// Mitsubishi GX Works2 project: ZhaoQing_OCV__Debug   PLC: Q10UDEH (continued)
     
     (*空框换内衬线体*)
    SwitchIO12203.xEntryEnable:=  ConveyorIO12125.xNextRun;
    ConveyorIO12142.iProductCategoryIn:=ConveyorIO12125.iProductCategoryOut;
    IF ConveyorIO12142.iProductCategory=4 THEN
    	SwitchIO12203.xSwithEnable:=1;
    ELSE
    	SwitchIO12203.xSwithEnable:=0;
    END_IF;
    SwitchIO12203.xExitEnable:=ConveyorIO12143.xEmpty;
    ConveyorIO12143.xLoad:=ConveyorIO12142.xNextRun;
    ConveyorIO12143.iProductCategoryIn:=ConveyorIO12142.iProductCategoryOut;
    ConveyorIO12143.xUnload:=ConveyorIO12144.xEmpty;
    (*OCV1线体*) 
  (*  ConveyorIO12144.xLoad:=ConveyorIO12143.xNextRun;*)
    SwitchIO12330.xEntryEnable:=ConveyorIO12143.xNextRun;
    ConveyorIO12144.iProductCategoryIn:=ConveyorIO12143.iProductCategoryOut;
    IF ConveyorIO12144.iProductCategory =2 THEN  (*临时程序  手动调试完毕后改为2*)
   	 SwitchIO12330.xSwithEnable:=1;
    ELSE
    SwitchIO12330.xSwithEnable:=0;	
    END_IF;   
    ConveyorIO12144.xUnload:=ConveyorIO12333.xEmpty AND SwitchIO12330.xSwithEnable=0;
     SwitchIO12330.xExitEnable:=ConveyorIO12160.xEmpty AND SwitchIO12330.xSwithEnable=1;
     ConveyorIO12160.xLoad:=Switch12330ConveyorOut.xNextRun;
     IF XA5 THEN(*人工按钮*)
     	IF ConveyorIO12146.xEmpty THEN
     		m_xOCV1Done:=1;
     	END_IF;
     	m_xPickOutDone :=1;
     END_IF;
     IF ConveyorIO12160.xEmpty THEN
     	m_xOCV1Done:=0;
     END_IF ;
     IF ConveyorIO12146.xEmpty THEN
     	m_xPickOutDone :=0;
     END_IF;
     ConveyorIO12160.tLoadDelay:=T#2s;
     ConveyorIO12160.xUnload:=ConveyorIO12146.xEmpty AND m_xOCV1Done;
     Y27F:=ConveyorIO12146.xEmpty AND m_xOCV1Done;(*阻挡气缸*)
     ConveyorIO12146.xLoad:= ConveyorIO12160.xNextRun;
     (*OCV2线体*)    
    SwitchIO12333.xEntryEnable:=ConveyorIO12144.xNextRun;
	SwitchIO12333.xSwithEnable:=1;
	SwitchIO12333.xExitEnable:=NOT XAE;
     (*空框换内衬线体*)    	
     SwitchIO12204.xEntryEnable:=1;
      SwitchIO12204.xSwithEnable:=1;
      SwitchIO12204.xExitEnable:=ConveyorIO12151.xEmpty;
      ConveyorIO12151.xLoad:=ConveyorIO12204.xNextRun;
      ConveyorIO12151.xUnload:=ConveyorIO12150.xEmpty;
      ConveyorIO12150.xLoad:=ConveyorIO12151.xNextRun;
      ConveyorIO12150.xUnload:=ConveyorIO12149.xEmpty;
      SwitchIO12328.xEntryEnable:=ConveyorIO12150.xNextRun;
       SwitchIO12328.xSwithEnable:=1;
	(****************提升机8******************)
	Lifter8Priority(xCondition1:= NOT ConveyorIO12148.xEmpty,
	                          xCondition2:= NOT ConveyorIO12146.xEmpty AND m_xPickOutDone  ,
	                          xCondition3:= FALSE,(*成品库车间空框回流线体不为空的条件*)
	                          xCondition4:= FALSE ,
	                          xCondition5:= FALSE ,
	                          xTaskComplete:= LDF(TRUE,Conveyor8IO.xEmpty=0) ,
	                          xReset:=g_xResetSingle AND g_iDeviceIDSelect=8,
	                          iPriority:= m_iLifter8Task);
	     D16:=m_iLifter8Task;(*触摸屏显示当前任务*)
		CASE m_iLifter8Task OF
			1:(*空框回流线体*)
				Lifter8IO.iDestinationPos:=2;
				SwitchIO12328.xExitEnable:=Lifter8IO.iCurrentPos=2 AND XC2 AND Conveyor8IO.xEmpty AND NOT XC1;
			   Conveyor8IO.xLoad:=ConveyorIO12148.xNextRun;
               Conveyor8IO.xloadCCW:=1;
			2:(*OCV1*)
				Lifter8IO.iDestinationPos:=1;
			   Conveyor8IO.xLoad:=ConveyorIO12146.xNextRun;
			   ConveyorIO12146.xUnload:=Conveyor8Io.xEmpty AND Lifter8IO.iCurrentPos=1 AND XC1 AND XC2;
			   Y27E:=Conveyor8Io.xEmpty AND Lifter8IO.iCurrentPos=1 AND XC1 AND XC2;(*分拣位置阻挡气缸*)
               Conveyor8IO.xloadCCW:=0;			
			3:(*成品库对接*)
				Lifter8IO.iDestinationPos:=4;
			(*	Conveyor8IO.xLoad:=ConveyorIO12147.xNextRun;*)
				Conveyor8IO.xloadCCW:=0;
				ELSE
				Conveyor8IO.xLoad:=0;
				SwitchIO12328.xExitEnable:=0;
				ConveyorIO12146.xUnload:=0;
				Y27E:=0;(*分拣位置阻挡气缸*)
		END_CASE;		
	IF Conveyor8IO.xEmpty=0 THEN
		Lifter8IO.xMDIExe:=1;
		Lifter8IO.iDestinationPos:=3;
	END_IF;	
	IF Lifter8IO.iCurrentPos=3 AND XC3 THEN
		Conveyor8Io.xUnload:=ConveyorIO12159.xEmpty;
		Conveyor8IO.xUnloadCCW:=1;
	ELSE
		Conveyor8Io.xUnload:=0;
	END_IF;	
	ConveyorIO12159.xLoad:=Conveyor8IO.xNextRun;
   ConveyorIO12159.xUnload:=ConveyorIO12158.xEmpty;
   SwitchIO12337.xEntryEnable:=ConveyorIO12159.xNextRun;
   SwitchIO12337.xSwithEnable:=1;
   SwitchIO12337.xLiftCylinderExtendInit:=1;
   SwitchIO12337.xExitEnable:=ConveyorIO12156.xEmpty;
   ConveyorIO12156.xLoad:=ConveyorIO12157.xNextRun;
	(**********常温库入库分流*******************)	
	ConveyorIO12156.xUnload:=ConveyorIO12155.xEmpty;
	ConveyorIO12155.xLoad:=ConveyorIO12156.xNextRun;
	     (*触摸屏上计数与清零程序*)
     IF LDF(TRUE,ConveyorIO12155.xEmpty) THEN
     	D14:=D14+1;
     END_IF;
     IF M169 THEN
     	D14:=0;
     END_IF;
	
	(**********常温库1巷道入库*******************) 
         	ConveyorIO12155.xUnload:=ConveyorIO12141.xEmpty AND ConveyorIO12155.iProductCategory>1 ;
         	ConveyorIO12141.xLoad:=ConveyorIO12155.xNextRun;
         	ConveyorIO12141.xUnload:=ConveyorIO12321.xEmpty;
            (*分流信息传递到巷道1的顶升移载处*)        	
  			ConveyorIO12141.iProductCategoryIn:= ConveyorIO12155.iProductCategoryOut;    
  			    
            SwitchIO12321.xEntryEnable:=ConveyorIO12141.xNextRun;
			ConveyorIO12321.iProductCategoryIn:=ConveyorIO12141.iProductCategoryOut;
           (*分流信息显示为本巷道，启动顶升移载*)
           IF ConveyorIO12321.iProductCategory=2 THEN
          	 SwitchIO12321.xSwithEnable:=1;
           ELSE
      	     	SwitchIO12321.xSwithEnable:=0;
           END_IF;
           (*双料入库，优先选择1 ，当1结束后恢复到0，2秒 ，然后再跳到2,0状态用来复位移载的出料*) 
          m_tonSwitch1NOSeleteDelay(IN:= m_iSwitch12321Select=0 ,PT:= t#2S ,Q:=m_xSwitch12321NoSeleteDelay,ET:= m_tSwitch12321NOSeleteCurrent);
         IF   m_xSwitch12321NoSeleteDelay THEN
         	m_xSwitch12321Select:=1;
         END_IF;
         IF ldf(TRUE,ConveyorIO12138.xEmpty)  OR ldf(TRUE,ConveyorIO12139.xEmpty) THEN
         	m_xSwitch12321Select:=0;
         END_IF;
           IF ConveyorIO12139.xEmpty AND  m_xSwitch12321Select  THEN
           		m_iSwitch12321Select:=1;
	           	ELSIF NOT ConveyorIO12139.xEmpty  AND ConveyorIO12138.xEmpty AND m_xSwitch12321Select THEN
           	  	m_iSwitch12321Select:=2;
          	 ELSE
           		m_iSwitch12321Select:=0;
           END_IF;
           IF SwitchIO12321.xSwithEnable THEN
         	  SwitchIO12321.xExitEnable:=((ConveyorIO12139.xEmpty AND m_iSwitch12321Select=1) 
                                                          OR   (ConveyorIO12138.xEmpty AND m_iSwitch12321Select=2)) AND CylinderIO12320.iCurrentPos=1;
           ELSE(*分流到下一巷道*)
   	        	 SwitchIO12321.xExitEnable:= ConveyorIO12137.xEmpty;
    	        ConveyorIO12137.xLoad:= ConveyorIO12321.xNextRun ;
    	         ConveyorIO12137.iProductCategoryIn:=   ConveyorIO12321.iProductCategoryOut;     
            END_IF;
 
           ConveyorIO12139.xLoad:=ConveyorIO12140.xNextRun AND m_iSwitch12321Select=1 ;
   	       ConveyorIO12138.xLoad:=ConveyorIO12140.xNextRun AND m_iSwitch12321Select=2 ;
   	       IF  ConveyorIO12138.xEmpty =0 AND ConveyorIO12139.xEmpty =0 AND X72 AND X74 THEN
   	       	CylinderIO12320.xMDIExe:=1;
   	       	CylinderIO12320.iDestinationPos:=2;
   	       	ConveyorIO12138.xPutInto:=0;
   	       	ConveyorIO12139.xPutInto:=0;
   	       END_IF;
   	       IF g_xImport1Force THEN (* 1巷道单框强制入库*)
   	       	CylinderIO12320.xMDIExe:=1;
   	       	CylinderIO12320.iDestinationPos:=2;
   	       	ConveyorIO12138.xPutInto:=0;
   	       	ConveyorIO12139.xPutInto:=0;   
   	       	END_IF;	       
   	       IF NOT X72 AND NOT X74 THEN
   	       		CylinderIO12320.xMDIExe:=1;
   	       		CylinderIO12320.iDestinationPos:=1;
   	       END_IF;
   	       IF LDP(TRUE,CylinderIO12320.iCurrentPos=1 AND NOT ConveyorIO12138.xCWPresent AND NOT ConveyorIO12139.xCWPresent) THEN   	       	
   	       		ConveyorIO12138.xPutInto:=1;
   	       		ConveyorIO12139.xPutInto:=1;
   	       END_IF;        
	(**********常温库2巷道入库*******************)
	       ConveyorIO12137.xUnload:=ConveyorIO12136.xEmpty;
	       ConveyorIO12136.xLoad:=ConveyorIO12137.xNextRun;	       
  		   ConveyorIO12136.iProductCategoryIn:= ConveyorIO12137.iProductCategoryOut;  
         	ConveyorIO12136.xUnload:=ConveyorIO12135.xEmpty AND ConveyorIO12136.iProductCategory>2 ;
            (*分流信息传递到巷道1的顶升移载处*)        	
  			ConveyorIO12135.iProductCategoryIn:= ConveyorIO12136.iProductCategoryOut;       			    
            SwitchIO12317.xEntryEnable:=ConveyorIO12136.xNextRun;
           (*分流信息显示为本巷道，启动顶升移载*)
           IF ConveyorIO12135.iProductCategory=3 THEN
          	 SwitchIO12317.xSwithEnable:=1;
           ELSE
      	     	SwitchIO12317.xSwithEnable:=0;
           END_IF;
           (*双料入库，优先选择1 ，当1结束后恢复到0，2秒 ，然后再跳到2,0状态用来复位移载的出料*) 
          m_tonSwitch2NOSeleteDelay(IN:= m_iSwitch12317Select=0 ,PT:= t#2S ,Q:=m_xSwitch12317NoSeleteDelay,ET:= m_tSwitch12317NOSeleteCurrent);
         IF   m_xSwitch12317NoSeleteDelay THEN
         	m_xSwitch12317Select:=1;
         END_IF;
         IF ldf(TRUE,ConveyorIO12132.xEmpty)  OR ldf(TRUE,ConveyorIO12133.xEmpty) THEN
         	m_xSwitch12317Select:=0;
         END_IF;
           IF ConveyorIO12133.xEmpty AND  m_xSwitch12317Select   THEN
           		m_iSwitch12317Select:=1;
	           	ELSIF NOT ConveyorIO12133.xEmpty  AND ConveyorIO12132.xEmpty AND m_xSwitch12317Select THEN
           	  	m_iSwitch12317Select:=2;
          	 ELSE
           		m_iSwitch12317Select:=0;
           END_IF;
           IF SwitchIO12317.xSwithEnable THEN
         	  SwitchIO12317.xExitEnable:=((ConveyorIO12133.xEmpty AND m_iSwitch12317Select=1) 
                                                          OR   (ConveyorIO12132.xEmpty AND m_iSwitch12317Select=2)) AND CylinderIO12316.iCurrentPos=1;
           ELSE(*分流到下一巷道*)
   	        	 SwitchIO12317.xExitEnable:= ConveyorIO12131.xEmpty;
    	        ConveyorIO12131.xLoad:= ConveyorIO12135.xNextRun ;
    	        ConveyorIO12131.iProductCategoryIn:=ConveyorIO12135.iProductCategoryOut;
            END_IF;
           	                                          
           ConveyorIO12133.xLoad:=ConveyorIO12134.xNextRun AND m_iSwitch12317Select=1 ;
   	       ConveyorIO12132.xLoad:=ConveyorIO12134.xNextRun AND m_iSwitch12317Select=2 ;
   	       IF  ConveyorIO12133.xEmpty =0 AND ConveyorIO12132.xEmpty =0 AND CylinderIO12316.xPresentDetect1 AND CylinderIO12316.xPresentDetect2 THEN
   	       	CylinderIO12316.xMDIExe:=1;
   	       	CylinderIO12316.iDestinationPos:=2;
   	       	ConveyorIO12133.xPutInto:=0;
   	       	ConveyorIO12132.xPutInto:=0;
   	       END_IF;
   	       IF g_xImport2Force THEN (* 1巷道单框强制入库*)
   	       	CylinderIO12316.xMDIExe:=1;
   	       	CylinderIO12316.iDestinationPos:=2;
   	       	ConveyorIO12133.xPutInto:=0;
   	       	ConveyorIO12132.xPutInto:=0;   
   	       	END_IF;	       
   	       IF NOT CylinderIO12316.xPresentDetect1 AND NOT CylinderIO12316.xPresentDetect2 THEN
   	       		CylinderIO12316.xMDIExe:=1;
   	       		CylinderIO12316.iDestinationPos:=1;
   	       END_IF;
   	       IF LDP(TRUE,CylinderIO12316.iCurrentPos=1 AND NOT ConveyorIO12132.xCWPresent AND NOT ConveyorIO12133.xCWPresent) THEN   	       	
   	       		ConveyorIO12133.xPutInto:=1;
   	       		ConveyorIO12132.xPutInto:=1;
   	       END_IF;  
	(**********常温库3巷道入库*******************)
	       ConveyorIO12131.xUnload:=ConveyorIO12130.xEmpty AND ConveyorIO12131.iProductCategory>3 ;
	       ConveyorIO12130.xLoad:=ConveyorIO12131.xNextRun;	       
  		   ConveyorIO12130.iProductCategoryIn:= ConveyorIO12131.iProductCategoryOut;  
            (*分流信息传递到巷道1的顶升移载处*)   
             ConveyorIO12130.xUnload:=ConveyorIO12129.xEmpty;
             SwitchIO12314.xEntryEnable:=ConveyorIO12130.xNextRun;   	
  			ConveyorIO12129.iProductCategoryIn:= ConveyorIO12130.iProductCategoryOut;       			               
           (*分流信息显示为本巷道，启动顶升移载*)
           IF ConveyorIO12129.iProductCategory=4THEN
          	 SwitchIO12314.xSwithEnable:=1;
           ELSE
      	     	SwitchIO12314.xSwithEnable:=0;
           END_IF;
           (*双料入库，优先选择1 ，当1结束后恢复到0，2秒 ，然后再跳到2,0状态用来复位移载的出料*) 
          m_tonSwitch3NOSeleteDelay(IN:= m_iSwitch12314Select=0 ,PT:= t#2S ,Q:=m_xSwitch12314NoSeleteDelay,ET:= m_tSwitch12314NOSeleteCurrent);
         IF   m_xSwitch12314NoSeleteDelay THEN
         	m_xSwitch12314Select:=1;
         END_IF;
         IF ldf(TRUE,ConveyorIO12126.xEmpty)  OR ldf(TRUE,ConveyorIO12127.xEmpty) THEN
         	m_xSwitch12314Select:=0;
         END_IF;
           IF ConveyorIO12127.xEmpty AND  m_xSwitch12314Select   THEN
           		m_iSwitch12314Select:=1;
	           	ELSIF NOT ConveyorIO12127.xEmpty  AND ConveyorIO12126.xEmpty AND m_xSwitch12314Select THEN
           	  	m_iSwitch12314Select:=2;
          	 ELSE
           		m_iSwitch12314Select:=0;
           END_IF;
           IF SwitchIO12314.xSwithEnable THEN
         	  SwitchIO12314.xExitEnable:=((ConveyorIO12127.xEmpty AND m_iSwitch12314Select=1) 
                                                          OR   (ConveyorIO12126.xEmpty AND m_iSwitch12314Select=2)) AND CylinderIO12313.iCurrentPos=1;
           ELSE(*分流到下一巷道*)
				;(*报警*)
            END_IF;
           	                                          
           ConveyorIO12127.xLoad:=ConveyorIO12128.xNextRun AND m_iSwitch12314Select=1 ;
   	       ConveyorIO12126.xLoad:=ConveyorIO12128.xNextRun AND m_iSwitch12314Select=2 ;
   	       IF  ConveyorIO12126.xEmpty =0 AND ConveyorIO12127.xEmpty =0 AND CylinderIO12313.xPresentDetect1 AND CylinderIO12313.xPresentDetect2 THEN
   	       	CylinderIO12313.xMDIExe:=1;
   	       	CylinderIO12313.iDestinationPos:=2;
   	       	ConveyorIO12126.xPutInto:=0;
   	       	ConveyorIO12127.xPutInto:=0;
   	       END_IF;
   	       IF g_xImport3Force THEN (* 1巷道单框强制入库*)
   	       	CylinderIO12313.xMDIExe:=1;
   	       	CylinderIO12313.iDestinationPos:=2;
   	       	ConveyorIO12126.xPutInto:=0;
   	       	ConveyorIO12127.xPutInto:=0;   
   	       	END_IF;	       
   	       IF NOT CylinderIO12313.xPresentDetect1 AND NOT CylinderIO12313.xPresentDetect2 THEN
   	       		CylinderIO12313.xMDIExe:=1;
   	       		CylinderIO12313.iDestinationPos:=1;
   	       END_IF;
   	       IF LDP(TRUE,CylinderIO12313.iCurrentPos=1 AND NOT ConveyorIO12127.xCWPresent AND NOT ConveyorIO12126.xCWPresent) THEN   	       	
   	       		ConveyorIO12126.xPutInto:=1;
   	       		ConveyorIO12127.xPutInto:=1;
   	       END_IF;  
END_IF;
(*人工操作按钮*)
IF LDP(TRUE,X0FF)  AND NOT  Y290 THEN
	 m_xMotorFlag:=1;
ELSE
	m_xMotorFlag:=0;
END_IF;

IF m_xMotorFlag THEN
	Y290:=1;
	Y27A:=1;
	Y27B:=1;
END_IF;

IF LDP(TRUE,X0FF) AND NOT m_xMotorFlag THEN
	Y290:=0;
	Y27A:=0;
	Y27B:=0;
END_IF;
(*报警*)
M500:=D2330=1;(*常温库出库分流读码失败*)
M501:=D2325=1;(*常温库入库分流读码失败*)
g_xAlarm:=M500 
                     OR M501;
END_PROGRAM

FUNCTION_BLOCK PriorityFB
VAR_INPUT
  xCondition1 : BOOL;  (* 条件1 *)
  xCondition2 : BOOL;  (* 条件2 *)
  xCondition3 : BOOL;  (* 条件3 *)
  xCondition4 : BOOL;  (* 条件4 *)
  xCondition5 : BOOL;  (* 条件5 *)
  xTaskComplete : BOOL;  (* 任务完成 *)
  xReset : BOOL;  (* 复位 *)
END_VAR
VAR
  xOccupy : BOOL;  (* 占用 *)
END_VAR
VAR_OUTPUT
  iPriority : INT;  (* 输出任务号 *)
END_VAR
VAR
  m_tonCondition1Delay : TON;
  m_xCondition1Delay : BOOL;
  m_tCondition1CurrentTime : TIME;
  arriTaskStack : ARRAY [0..5] OF INT;
  m_tonCondition2Delay : TON;
  m_xCondition2Delay : BOOL;
  m_tCondition2CurrentTime : TIME;
  m_tonCondition3Delay : TON;
  m_xCondition3Delay : BOOL;
  m_tCondition3CurrentTime : TIME;
  m_tonCondition4Delay : TON;
  m_xCondition4Delay : BOOL;
  m_tCondition4CurrentTime : TIME;
  m_tonCondition5Delay : TON;
  m_xCondition5Delay : BOOL;
  m_tCondition5CurrentTime : TIME;
  jj : INT;
END_VAR
(****************************************************************************)
(*
优先级功能块，存储5个条件的优先级，实现栈功能先入先出，
复位功能还有问题，
*)
(***************************************************************************)
m_tonCondition1Delay(IN:= xCondition1 AND NOT xReset ,PT:= T#1s,Q:= m_xCondition1Delay , ET:= m_tCondition1CurrentTime );
m_tonCondition2Delay(IN:= xCondition2 AND NOT xReset ,PT:= T#1s,Q:= m_xCondition2Delay , ET:= m_tCondition2CurrentTime );
m_tonCondition3Delay(IN:= xCondition3 AND NOT xReset ,PT:= T#1s,Q:= m_xCondition3Delay , ET:= m_tCondition3CurrentTime );
m_tonCondition4Delay(IN:= xCondition4 AND NOT xReset ,PT:= T#1s,Q:= m_xCondition4Delay , ET:= m_tCondition4CurrentTime );
m_tonCondition5Delay(IN:= xCondition5 AND NOT xReset ,PT:= T#1s,Q:= m_xCondition5Delay , ET:= m_tCondition5CurrentTime );

IF ldp(TRUE,m_xCondition1Delay) THEN
	FOR jj:=0 TO 5 BY 1 DO
		IF arriTaskStack[jj]=0 THEN
			arriTaskStack[jj]:=1;
			EXIT;
		END_IF;		
	END_FOR;
END_IF;

IF ldp(TRUE,m_xCondition2Delay) THEN
	FOR jj:=0 TO 5 BY 1 DO
		IF arriTaskStack[jj]=0 THEN
			arriTaskStack[jj]:=2;
			EXIT;
		END_IF;		
	END_FOR;
END_IF;

IF ldp(TRUE,m_xCondition3Delay) THEN
	FOR jj:=0 TO 5 BY 1 DO
		IF arriTaskStack[jj]=0 THEN
			arriTaskStack[jj]:=3;
			EXIT;
		END_IF;		
	END_FOR;
END_IF;

IF ldp(TRUE,m_xCondition4Delay) THEN
	FOR jj:=0 TO 5 BY 1 DO
		IF arriTaskStack[jj]=0 THEN
			arriTaskStack[jj]:=4;
			EXIT;
		END_IF;		
	END_FOR;
END_IF;

IF ldp(TRUE,m_xCondition5Delay) THEN
	FOR jj:=0 TO 5 BY 1 DO
		IF arriTaskStack[jj]=0 THEN
			arriTaskStack[jj]:=5;
			EXIT;
		END_IF;		
	END_FOR;
END_IF;

iPriority:=arriTaskStack[0];

IF 	LDP(TRUE, xTaskComplete) THEN
	FOR jj:=0 TO 4 BY 1 DO
		arriTaskStack[jj]:=arriTaskStack[jj+1];
	END_FOR;
		arriTaskStack[5]:=0;
END_IF;

IF LDP(TRUE,xReset) THEN
		FOR jj:=0 TO 5 BY 1 DO
		arriTaskStack[jj]:=0;
	END_FOR;
END_IF;
END_FUNCTION_BLOCK

FUNCTION ShuttleCarCurrentPosition
VAR_INPUT
  xPosition1 : BOOL;
  xPosition2 : BOOL;
  xPosition3 : BOOL;
END_VAR
(************************************
计算输送车当前位置的函数
**************************************)
IF xPosition1 THEN
	ShuttleCarCurrentPosition:=1;
END_IF;
IF xPosition2 THEN
	ShuttleCarCurrentPosition:=2;
END_IF;
IF xPosition3 THEN
	ShuttleCarCurrentPosition:=3;
END_IF;
END_FUNCTION

FUNCTION ShuttleCarVelocityEncoder
VAR_INPUT
  iDestinationPos : INT;  (* 目标位置 *)
  iCurrentPos : INT;  (* 当前位置 *)
  xEnable : BOOL;  (* 使能 *)
END_VAR
IF xEnable THEN
	IF ABS(iCurrentPos-iDestinationPos)<300  THEN
		ShuttleCarVelocityEncoder:=0;
	ELSE
		ShuttleCarVelocityEncoder:=1;
	END_IF;
ELSE
	ShuttleCarVelocityEncoder:=0;
END_IF;
END_FUNCTION

FUNCTION_BLOCK ShuttleCarVelocityFB
VAR_INPUT
  xEnable : BOOL;  (* 使能 *)
  xMotorCW : BOOL;  (* 电机正转 *)
  xMotorCCW : BOOL;  (* 电机反转 *)
  xPosition1Switch : BOOL;  (* 位置1开关 *)
  xDecelerationSwitch : BOOL;  (* 减速开关 *)
  xPosition2Switch : BOOL;  (* 位置2开关 *)
END_VAR
VAR
  iFloor : INT;  (* 层数 *)
END_VAR
VAR_OUTPUT
  xHighSpeed : BOOL;
END_VAR
IF xEnable THEN
	(*电机旋转，并且在位置开关上的时候触发加速*)
	IF( LDP(TRUE,xMotorCW) AND xPosition1Switch ) OR (  LDP(TRUE,xMotorCCW) AND xPosition2Switch) THEN
		xHighSpeed:=1;
		iFloor:=0;
	END_IF;
	IF LDF(TRUE,xMotorCW) OR LDF(TRUE,xMotorCCW) THEN
		xHighSpeed:=0;
    END_IF;
	IF LDP(TRUE,xDecelerationSwitch) THEN
		iFloor:=iFloor+1;
	END_IF;
	IF iFloor=2 THEN
		xHighSpeed:=0;
		iFloor:=0;
	END_IF;
ELSE
    xHighSpeed:=0;
END_IF;
END_FUNCTION_BLOCK

PROGRAM Start
IF g_xReset THEN
	SM50:=1;
ELSE
	SM50:=0;
END_IF;
CASE g_iState OF
	0: 
		g_xManual:=1;
		g_xAuto:=0;	
		g_xStackLampAmber:=1;
		g_xStackLampGreen:=0;
		g_xRemoteAuto:=0;
	1:
		g_xManual:=0;
		g_xAuto:=1;
		g_xStackLampGreen:=1;
		g_xStackLampAmber:=0;
		g_xRemoteAuto:=0;
	2:	
        g_xRemoteAuto:=1;
        g_xStackLampGreen:=1;
        g_xStackLampAmber:=0;
        g_xAuto:=0;
		g_xManual:=0;
END_CASE;
IF g_xLocalAutoStart THEN  
	g_iState:=1;
END_IF;
IF g_xAlarm AND SM412 THEN
	g_xStackLampRed:=1;
	g_xBuzzer:=1;
ELSE
	g_xStackLampRed:=0;
	g_xBuzzer:=0;	
END_IF;
IF g_xStop OR g_xEStop=0 THEN 
	g_iState:=0;
END_IF;
IF g_xRemoteAutoStart THEN
	g_iState:=2;
END_IF;
IF g_xPause AND SM412 THEN
	g_xStackLampGreen:=0;
	g_xStackLampAmber:=0;
END_IF;
END_PROGRAM

FUNCTION_BLOCK Switch
VAR_IN_OUT
  ConveyorEntryIO : ConveyorIO;
END_VAR
VAR
  ConveyorEntry : Conveyor;
END_VAR
VAR_IN_OUT
  ConveyorExitIO : ConveyorIO;
END_VAR
VAR
  m_tonLiftCylinderDelay : TON;  (* 顶升延时 *)
  m_xLiftCylinderDelay : BOOL;
  m_tLiftCylinderDelay : TIME;
  m_tonExitBarDelay : TON;  (* 退出阻挡器延时 *)
  m_tExitBarDelay : TIME;
  m_xExitBarDelay : BOOL;
END_VAR
VAR_IN_OUT
  SwitchIO : SwitchIO;
END_VAR
VAR
  iStep : INT;
  ConveyorExit : Conveyor;
  m_xInitial : BOOL;
  m_tonCylinderOvertime : TON;  (* 气缸超时报警定时器 *)
  m_tCylinderOvertimeCurrent : TIME;
END_VAR
(**************************************************
顶升移载模块，抽象为一条输入输线 ，一条输出输送线
一个进入阻挡器，一个放出阻挡器，和一个顶升气缸的控制
程序思路比较混乱，接口不清晰，需要整改
直接放行的时候有问题
switchEnable =0的时候   离开线体的PutInto有问题
增加xPutInto程序
12-17日   V1.0
***************************************************)
ConveyorEntry(ConveyorMotor:=ConveyorEntryIO);
ConveyorExit(ConveyorMotor:=ConveyorExitIO);


IF NOT m_xInitial THEN
	
	m_xInitial:=1;
END_IF;
IF g_xAuto THEN
	CASE iStep OF
		0:(*初始化*)
		ConveyorEntryIO.xLoad:=0;
		ConveyorEntryIO.xUnload:=0;
		ConveyorEntryIO.xPutInto:=0;
		ConveyorExitIO.xLoad:=0;
		ConveyorExitIo.xUnload:=0;
		ConveyorExitIO.xPutInto:=0;
		SwitchIO.xEntryBarCylinderRetract:=0;
		SwitchIO.xExitBarCylinderRetract:=0;
		IF SwitchIO.xLiftCylinderExtendInit THEN
			SwitchIO.xLiftCylinderExtend:=1;
			SwitchIO.xLiftCylinderRetract:=0;
		    IF SwitchIO.xLiftCylinderExtendDetect THEN
			    iStep:=1;
		     END_IF; 
		ELSE
			SwitchIO.xLiftCylinderExtend:=0;
			SwitchIO.xLiftCylinderRetract:=1;	
		    IF SwitchIO.xLiftCylinderRetractDetect THEN
			    iStep:=1;
		    END_IF;		
		END_IF;
		1:(*上料*)
        IF SwitchIO.xEntryEnable AND ConveyorEntryIO.xEmpty AND ConveyorExitIO.xEmpty THEN
        	SwitchIO.xEntryBarCylinderRetract:=1;
        	ConveyorEntryIO.xLoad:=1;
        END_IF;
        IF ConveyorEntryIO.xEmpty=0 THEN
        	SwitchIO.xEntryBarCylinderRetract:=0;
        	ConveyorEntryIO.xLoad:=0;
        	ConveyorExitIO.xPutInto:=1;
        END_IF;
        IF m_xLiftCylinderDelay AND  SwitchIO.xSwithEnable THEN
        	 iStep:=2;
        END_IF;
        IF SwitchIO.xSwithEnable=0 AND m_xLiftCylinderDelay  THEN
        	 iStep:=3;
        END_IF;
		2:(*顶升*)
		   ConveyorExitIO.iProductCategory:=ConveyorEntryIO.iProductCategory;
			SwitchIO.xExitBarCylinderRetract:=0;
		    IF SwitchIO.xLiftCylinderExtendInit THEN
			    SwitchIO.xLiftCylinderExtend:=0;
			    SwitchIO.xLiftCylinderRetract:=1;
		    ELSE
			    SwitchIO.xLiftCylinderExtend:=1;
			    SwitchIO.xLiftCylinderRetract:=0;			
		   END_IF;

		  IF SwitchIO.xLiftCylinderExtendInit THEN
		  	IF SwitchIO.xLiftCylinderRetractDetect THEN
		  		iStep:=4;
		  	END_IF;
		  	ELSE
		  	IF SwitchIO.xLiftCylinderExtendDetect THEN
		      iStep:=4; 
		  	END_IF;
		  END_IF;
		  3:(*放行*)	
		    ConveyorExitIO.iProductCategory:=ConveyorEntryIO.iProductCategory;
		  	SwitchIO.xExitBarCylinderRetract:=1;
		  	ConveyorExitIO.xPutInto:=0;
		  	iStep:=4;
		  4:(*下料*)
		  (*通过出料传输线下料*)
		  IF SwitchIO.xExitEnable  AND m_xExitBarDelay AND NOT SwitchIO.xExitBarCylinderRetract  THEN		  
		  	ConveyorExitIO.xUnload:=1;
		  ELSE
		  	ConveyorExitIO.xUnload:=0;
		  END_IF;	
		   (*通过进料传输线下料*)
		  IF SwitchIO.xExitEnable  AND m_xExitBarDelay  AND SwitchIO.xExitBarCylinderRetract THEN		  
		  	ConveyorEntryIO.xUnload:=1;
		  ELSE
		  	ConveyorEntryIO.xUnload:=0;
		  END_IF;			    	
		  IF (ConveyorExitIO.xEmpty OR ConveyorEntryIO.xEmpty) AND m_xExitBarDelay  THEN
		  	ConveyorExitIO.xPutInto:=1;
		  	ConveyorEntryIO.xPutInto:=1;
			iStep:=0; 
		  END_IF;
	END_CASE;
        m_tonLiftCylinderDelay(IN:=NOT ConveyorEntryIO.xEmpty AND iStep=1 ,PT:= T#1S ,Q:= m_xLiftCylinderDelay ,ET:=m_tLiftCylinderDelay );
 		m_tonExitBarDelay(IN:=iStep=4 ,PT:= T#1s ,Q:= m_xExitBarDelay ,ET:= m_tExitBarDelay);
END_IF;
(*复位程序*)
IF (g_xResetSingle AND  (g_iDeviceIDSelect=ConveyorEntryIO.iDeviceID OR g_iDeviceIDSelect=ConveyorExitIO.iDeviceID))
	OR LDP(TRUE,SwitchIO.xLiftCylinderExtendInit) 
	OR LDF(TRUE,SwitchIO.xLiftCylinderExtendInit) 
	OR LDP(TRUE,SwitchIO.xPutInto)  THEN
	ConveyorEntryIO.xPutInto:=1;
	ConveyorExitIO.xPutInto:=1;
	iStep:=0;
END_IF;

IF g_xManual  THEN
	iStep:=0;
	ConveyorEntryIO.xLoad:=0;
    ConveyorEntryIO.xUnload:=0;
	ConveyorEntryIO.xPutInto:=0;
	ConveyorExitIO.xLoad:=0;
	ConveyorExitIo.xUnload:=0;
	ConveyorExitIO.xPutInto:=0;
	SwitchIO.xEntryBarCylinderRetract:=0;
	SwitchIO.xExitBarCylinderRetract:=0;
	IF SwitchIO.xEntryBarCylinderRetractButton THEN
		SwitchIO.xEntryBarCylinderRetract:=1;
	ELSE
		SwitchIO.xEntryBarCylinderRetract:=0;
	END_IF;
		IF SwitchIO.xExitBarCylinderRetractButton THEN
		SwitchIO.xExitBarCylinderRetract:=1;
	ELSE
		SwitchIO.xExitBarCylinderRetract:=0;
		END_IF;
		IF SwitchIO.xLiftCylinderExtendButton AND NOT SwitchIO.xLiftCylinderRetractButton THEN
			SwitchIO.xLiftCylinderExtend:=1;
			SwitchIO.xLiftCylinderRetract:=0;
		END_IF;
		IF NOT SwitchIO.xLiftCylinderExtendButton AND  SwitchIO.xLiftCylinderRetractButton THEN
			SwitchIO.xLiftCylinderExtend:=0;
			SwitchIO.xLiftCylinderRetract:=1;
		END_IF;		 
END_IF;
(*气缸超时报警*)
m_tonCylinderOvertime(IN:= (SwitchIO.xLiftCylinderExtend AND NOT SwitchIO.xLiftCylinderExtendDetect) 
                                                OR  (SwitchIO.xLiftCylinderRetract AND NOT SwitchIO.xLiftCylinderRetractDetect) ,
                                               PT:= SwitchIO.tSetOvertime ,Q:= SwitchIO.xOvertimeAlarm ,ET:= m_tCylinderOvertimeCurrent );
END_FUNCTION_BLOCK

FUNCTION_BLOCK BarCylinder
VAR_IN_OUT
  BarCylinderIO : BarCylinderIO;
END_VAR
VAR
  m_xInitial : BOOL;  (* 初始化 *)
  m_tonLoadDelay : TON;  (* 上料延时 *)
  m_xLoadDelay : BOOL;  (* 上料延时标志位 *)
  m_tLoadDelayCurrentTime : TIME;  (* 上料延时当前时间 *)
END_VAR
  (***********************************************************************
阻挡器模块，
由一个行程开关，一个阻挡器，一个倍速链输送电机组成
具有手动与自动模式
xEmpty显示当前为空料的状态
xUnload为卸料信号，连接下一设备的xEmpty信号
*************************************************************************)

IF NOT m_xInitial THEN
	BarCylinderIO.tLoadDelay:=T#5s;
	m_xInitial:=1;
END_IF;
IF g_xManual THEN    (*手动*)
	BarCylinderIO.xNextRun:=0;
	IF BarCylinderIO.xBarCylinderButton THEN
		BarCylinderIO.xBarCylinder:=1;
	ELSE
		BarCylinderIO.xBarCylinder:=0;
	END_IF;
	IF BarCylinderIO.xTransportMotorCWButton 
		AND NOT BarCylinderIO.xTransportMotorCCWButton 
		AND NOT BarCylinderIO.xTransportMotorCCW   THEN
		BarCylinderIO.xTransportMotorCW:=1;
	ELSE
		BarCylinderIO.xTransportMotorCW:=0;
	END_IF;
	IF BarCylinderIO.xTransportMotorCCWButton 
		AND NOT BarCylinderIO.xTransportMotorCWButton 
		AND NOT BarCylinderIO.xTransportMotorCW   THEN
		BarCylinderIO.xTransportMotorCCW:=1;
	ELSE
		BarCylinderIO.xTransportMotorCCW:=0;
	END_IF;
END_IF;
IF g_xAuto THEN(*自动*)
    IF BarCylinderIO.xUnload  AND NOT BarCylinderIO.xEmpty AND NOT BarCylinderIO.xNextRun THEN(*收到卸料命令，当阻挡器不为空时*)
    	BarCylinderIO.xBarCylinder:=1;
    	BarCylinderIO.xNextRun:=1;(*确保下料命令只执行一次，防止物料在输送过程中又有卸料命令导致多次卸料*)
    	BarCylinderIO.xTransportMotorCW:=1;
    END_IF;
    IF NOT  BarCylinderIO.xUnload  THEN
    	BarCylinderIO.xNextRun:=0;
    	BarCylinderIO.xBarCylinder:=0;
    END_IF;
    m_tonLoadDelay(IN:= BarCylinderIO.xPresentSwitch ,PT:= BarCylinderIO.tLoadDelay ,Q:= m_xLoadDelay,ET:= m_tLoadDelayCurrentTime );
    IF m_xLoadDelay OR  BarCylinderIO.xNextRun  THEN
    	BarCylinderIO.xEmpty:=0;
    ELSE
    	BarCylinderIO.xEmpty:=1;
    END_IF;
    (*如果为空，气缸顶起*)
   IF  BarCylinderIO.xEmpty  THEN
   	   BarCylinderIO.xBarCylinder:=0;
   END_IF;
   	IF BarCylinderIO.xLoad AND BarCylinderIO.xEmpty  THEN
		BarCylinderIO.xTransportMotorCW:=1;
   	END_IF;  
   	IF (BarCylinderIO.xLoad=0 OR BarCylinderIO.xEmpty=0)  AND (BarCylinderIO.xUnload=0 OR BarCylinderIO.xEmpty) THEN
   		BarCylinderIO.xTransportMotorCW:=0;
   	END_IF;
END_IF;  
IF BarCylinderIO.xEmpty AND BarCylinderIO.xLoad=0 THEN
	BarCylinderIO.iProductCategory:=0;
END_IF;

IF NOT g_xEStop THEN
	 BarCylinderIO.xTransportMotorCW:=0;
	 BarCylinderIO.xTransportMotorCCW:=0;
	 BarCylinderIO.xBarCylinder:=0;
END_IF;
END_FUNCTION_BLOCK

FUNCTION_BLOCK ShuttleCar
VAR_IN_OUT
  ShuttleCarInOut : ShuttleCarIO;
END_VAR
VAR
  m_tonBrakeDelay : TON;  (* 延时 *)
  m_tBrakeDelayCurrentTime : TIME;
  m_tonArriveDelay : TON;  (* 到达延时计时器 *)
  m_xArriveDelay : BOOL;  (* 到达延时 *)
  m_tArriveDelayCurrentTime : TIME;  (* 到达延时当前时间 *)
  m_xInit : BOOL;  (* 初始化标志位 *)
  m_tonPauseDelay : TON;  (* 暂停减速 *)
  m_tPauseDelayCurrentTime : TIME;  (* 暂停延时当前时间 *)
  m_tonOvertimeAlarm : TON;  (* 超时报警定时器 *)
  m_tOvertimeCurrentTime : TIME;  (* 超时报警当前时间 *)
END_VAR
(*******************************************************************
输送小车程序，可用于使用认址片控制位置的输送车程序，可用于控制提升机，
使用了限位捕捉程序防止小车惯性过大冲过限位后继续行走，捕捉程序采用反
转复位，这样设计有弊端可能反转复位后车的位置并没有回到限位以内,当两个
限位同时碰到的时候，会使运料小车进入死锁状态，通过xPassLimit来解开死锁，
可以在触摸屏中使用一个带权限的按钮来进行控制，配合ShuttleCarCurrentPos
函数来计算位置信息
增加自动开始后将当前位置置为零的信号防止设备停在两个位置开关的中间
修改信息  修改后请增加版本
2018-1-22增加到位延时：到位延时时间可以设置，适应双向到位的位置开关，通过调整延时时间让穿梭车停在到位开关的中间
增加气缸控制信号
增加抱闸延时
增加超时报警
YAO      V1.0
2018-1-22 YAO V1.1
接口说明：
输入：
xReady    准备就绪信号，接变频器的准备就绪，无准备就绪信号的设备常置1
xForward   手动 正转
xBackward 手动 反转
iCurrentPos 当前位置信息，由外部函数给出
iDestinationPos  目标位置，自动情况下判断目标位置和当前位置的差，选择前进或后退
xPosLimit 正方向限位  常闭信号
xNegLimit 反方向限位  常闭信号
xMDIExe   自动行走使能
xPassLimit 限位屏蔽
tArriveDelay 到位延时时间设置，当前位置等于目标位置后延时相应时间后停止，默认为0
xCylinder 如果是气缸的把这个标志位置为1，
tBrakeDelay 打开抱闸延时，默认100ms。行走后会延时相应的时间打开抱闸，防止提升轴的掉落
xLooseDetect 松绳检测开关
输出：
xCW 正转输出
xCCW 反转输出
xBrake 抱闸输出 
xMDIDone 自动行走完成信号
xPosLimitCatch 正限位报警
xNegLimitCatch 负限位报警
xBusy 工作中信号
xLooseAlarm 松绳报警，报警后不可以下降，提升后如果没有松绳检测开关后复位报警信号


********************************************************************)
IF NOT m_xInit THEN
	ShuttleCarInOut.tArriveDelay:=T#0s;   (*到位延时初始化为0*)
	ShuttleCarInOut.tBrakeDelay:=T#100ms;(*抱闸延时初始化为100ms*)
	ShuttleCarInOut.tSetOverTime:=T#60s;(*超时报警初始化为1分钟*)
	m_xInit:=1;
END_IF;
(*如果是气缸的话屏蔽限位和Ready信号*)
IF ShuttleCarInOut.xCylinder THEN
	ShuttleCarInOut.xPosLimit:=1;
	ShuttleCarInOut.xNegLimit:=1;
	ShuttleCarInOut.xReady:=1;
END_IF;
(*限位捕捉，防止冲过限位开关，反转后复位*)
ShuttleCarInOut.xPosLimitCatch:=LDF(TRUE,ShuttleCarInOut.xPosLimit) OR ShuttleCarInOut.xPosLimitCatch;
IF ShuttleCarInOut.xCCW THEN  
	ShuttleCarInOut.xPosLimitCatch:=0;
END_IF;

ShuttleCarInOut.xNegLimitCatch:=LDF(TRUE,ShuttleCarInOut.xNegLimit) OR ShuttleCarInOut.xNegLimitCatch;
(*松绳报警*)
IF LDP(TRUE,ShuttleCarInOut.xLooseDetect) THEN	
	ShuttleCarInOut.xLooseAlarm:=1;
END_IF;
(*提升复位报警*)
IF ShuttleCarInOut.xCW AND NOT  ShuttleCarInOut.xLooseDetect THEN   
	ShuttleCarInOut.xLooseAlarm:=0; 
END_IF;

IF ShuttleCarInOut.xCW THEN   
	ShuttleCarInOut.xNegLimitCatch:=0; 
END_IF;

IF ShuttleCarInOut.xPassLimit OR
	g_xReset OR   (*增加复位按钮*)
	(ShuttleCarInOut.xNegLimitCatch 
	AND ShuttleCarInOut.xPosLimitCatch)  THEN  
	ShuttleCarInOut.xNegLimitCatch:=0; 
	ShuttleCarInOut.xPosLimitCatch:=0;
	ShuttleCarInOut.xLooseAlarm:=0;
END_IF;
IF ShuttleCarInOut.xReady AND g_xEStop THEN
(*手动*)
    IF g_xManual THEN  
	    IF ShuttleCarInOut.xForward 
			AND ShuttleCarInOut.xBackward=0 
			AND ShuttleCarInOut.xCCW=0 
			AND ShuttleCarInOut.xPosLimitCatch=0  THEN
		    ShuttleCarInOut.xCW:=1;
		    ELSE
		    ShuttleCarInOut.xCW:=0;
	    END_IF;
	    IF ShuttleCarInOut.xBackward 
			AND ShuttleCarInOut.xForward=0 
			AND ShuttleCarInOut.xCW=0 
			AND ShuttleCarInOut.xNegLimitCatch=0 
			AND ShuttleCarInOut.xLooseAlarm=0
			AND G_xEStop THEN  
		    ShuttleCarInOut.xCCW:=1;
		    ELSE
		    ShuttleCarInOut.xCCW:=0;
	    END_IF;
    END_IF;
    (**********)
(*自动*)
  IF g_xAuto  THEN  
  	(*点动*)
 		IF LDP(TRUE,ShuttleCarInOut.xForward) THEN
 			ShuttleCarInOut.xMDIExe:=1;
			ShuttleCarInOut.iDestinationPos:=ShuttleCarInOut.iCurrentPos+1;
		END_IF;
		IF LDP(TRUE,ShuttleCarInOut.xBackward) THEN
			ShuttleCarInOut.xMDIExe:=1;
			ShuttleCarInOut.iDestinationPos:=ShuttleCarInOut.iCurrentPos-1;
		END_IF;	 
	(*>>>>>>>>>>>>>>>>>>>>>>>>>>>>>>>>>>>>>*)	
	  IF ShuttleCarInOut.xMDIExe AND ShuttleCarInOut.iDestinationPos<>0 THEN	
	    IF ShuttleCarInOut.iCurrentPos<ShuttleCarInOut.iDestinationPos AND ShuttleCarInOut.xPosLimitCatch=0 THEN   (*正转*)
			ShuttleCarInOut.xCW:=1;
			ShuttleCarInOut.xCCW:=0;
			ShuttleCarInOut.xMDIDone:=0;
		END_IF;

		IF ShuttleCarInOut.iCurrentPos>ShuttleCarInOut.iDestinationPos AND ShuttleCarInOut.xNegLimitCatch=0 AND ShuttleCarInOut.xLooseAlarm=0 THEN   (*反转*)
			ShuttleCarInOut.xCCW:=1;
			ShuttleCarInOut.xCW:=0;
			ShuttleCarInOut.xMDIDone:=0;
		END_IF;
	m_tonArriveDelay(IN:= ShuttleCarInOut.iCurrentPos=ShuttleCarInOut.iDestinationPos ,
	                                    PT:= ShuttleCarInOut.tArriveDelay ,
	                                    Q:= m_xArriveDelay ,
	                                    ET:= m_tArriveDelayCurrentTime);
	     (*到位延时时间可以设置，适应双向到位的位置开关，通过调整延时时间让穿梭车停在到位开关的中间*)
		IF m_xArriveDelay AND NOT ShuttleCarInOut.xCylinder THEN
			ShuttleCarInOut.xCW:=0;
			ShuttleCarInOut.xCCW:=0;
			ShuttleCarInOut.xMDIDone:=1;
			ELSE
			ShuttleCarInOut.xMDIDone:=0;
		END_IF;

		IF ShuttleCarInOut.xPosLimitCatch THEN
			ShuttleCarInOut.xCW:=0;
			ShuttleCarInOut.xMDIDone:=0;
		END_IF;

		IF ShuttleCarInOut.xNegLimitCatch THEN
			ShuttleCarInOut.xCCW:=0;
			ShuttleCarInOut.xMDIDone:=0;
		END_IF;
		ELSE
		ShuttleCarInOut.xCW:=0;
		ShuttleCarInOut.xCCW:=0;
		ShuttleCarInOut.xMDIDone:=0;
	  END_IF;
	END_IF;
	ELSE  (*无就绪信号   或急停的情况下*)
		ShuttleCarInOut.xCW:=0;
		ShuttleCarInOut.xCCW:=0;	
END_IF;
    (*抱闸延时*)
m_tonBrakeDelay(IN:= ShuttleCarInOut.xCW OR ShuttleCarInOut.xCCW,
                                    PT:= ShuttleCarInOut.tBrakeDelay,
                                    Q:=ShuttleCarInOut.xBrake ,
                                    ET:= m_tBrakeDelayCurrentTime);

(*自动上电后把当前位置清零，防止穿梭车不在开关位置*)
IF LDP(TRUE,g_xAuto) THEN
	ShuttleCarInOut.iCurrentPos:=0;
END_IF;
IF ShuttleCarInOut.xCW OR ShuttleCarInOut.xCCW THEN
	ShuttleCarInOut.xBusy:=1;
	ELSE
	ShuttleCarInout.xBusy:=0;
END_IF;

(*暂停，带延时减速斜坡，ShuttleCarInOut.xPauseRamp为减速斜坡输出位*)
m_tonPauseDelay(IN:=g_xPause,PT:= T#2s ,Q:=ShuttleCarInOut.xPauseRamp,ET:= m_tPauseDelayCurrentTime );
IF ShuttleCarInOut.xPauseRamp THEN
	ShuttleCarInOut.xCW:=0;
	ShuttleCarInOut.xCCW:=0;
	ShuttleCarInOut.xBrake:=0;
END_IF;
(*超时报警*)
m_tonOvertimeAlarm(IN:= ShuttleCarInOut.xMDIExe AND (ShuttleCarInOut.iCurrentPos<>ShuttleCarInOut.iDestinationPos) ,
                                           PT:= ShuttleCarInOut.tSetOverTime,
                                           Q:= ShuttleCarInOut.xOvertimeAlarm ,
                                           ET:= m_tOvertimeCurrentTime );
END_FUNCTION_BLOCK
